// TIA Portal project "SSA-3GHz_V18" (V18)

(* hardware
DEVICE "S7-1200"  S7-1200 Station
   slot 0: "Stand.sectionalRail35mmLength483mm_0"  S7-1200 Rack  Rack  V1.0
   slot 1: "S7-1200"  CPU 1215C DC/DC/DC  6ES7 215-1AG40-0XB0  V4.5
   slot 2: "AnalogInputSM12314AI_2"  6ES7 231-4HD32-0XB0  V2.0
   slot 3: "S7-1200analogInputSM1231RTD4AI_3"  SM 1231 AI4 x RTD  6ES7 231-5PD32-0XB0  V2.0
DEVICE "HMI_1"  KTP400 Basic PN
   slot 0: "HMI_1"  KTP400 Basic PN  6AV2 123-2DB03-0AX0  15.1.0.0
   slot 1: "HMI_RT_1"  KTP400 Basic PN  6AV2 123-2DB03-0AX0  15.1.0.0
   slot 5: "HMI_1.IE_CP_1"  PROFINET Interface  15.0.1.0
      slot 1: "PROFINET Interface_1"  PROFINET Interface
         slot 1: "Port_1"  Port
*)

// ===== PLC "S7-1200"  CPU 1215C DC/DC/DC =====

VAR_GLOBAL   // PLC tag table "Default tag table"
   "System_Byte" AT %MB1 : Byte;
   "FirstScan" AT %M1.0 : Bool;
   "DiagStatusUpdate" AT %M1.1 : Bool;
   "AlwaysTRUE" AT %M1.2 : Bool;
   "AlwaysFALSE" AT %M1.3 : Bool;
   "Clock_Byte" AT %MB0 : Byte;
   "Clock_10Hz" AT %M0.0 : Bool;
   "Clock_5Hz" AT %M0.1 : Bool;
   "Clock_2.5Hz" AT %M0.2 : Bool;
   "Clock_2Hz" AT %M0.3 : Bool;
   "Clock_1.25Hz" AT %M0.4 : Bool;
   "Clock_1Hz" AT %M0.5 : Bool;
   "Clock_0.625Hz" AT %M0.6 : Bool;
   "Clock_0.5Hz" AT %M0.7 : Bool;
   "MoveBlkStat" AT %MW100 : Int;
   "tmp_setIP" AT %I1.1 : Bool;
   "Tag_2" AT %I1.2 : Bool;
   "Pulse_mem" AT %M10.1 : Bool;
   "Tag_3" AT %Q1.1 : Bool;
   "Modbus_srv_enable" AT %M2.3 : Bool;   // ModBus Server Enable bit
END_VAR

VAR_GLOBAL   // PLC tag table "Test tags"
   "Counter" AT %MD100 : UDInt;
   "TestBlink" AT %Q1.0 : Bool;
   "VisuTest" AT %MB104 : Byte;
   "Set_IP_PArameters" AT %M10.2 : Bool;
END_VAR

VAR_GLOBAL   // PLC tag table "Analog I/O"
   "U_drain_RBK" AT %IW64 : Int;   // Drain voltage read-back
   "U_drain" AT %QW64 : Int;   // Drain voltage set-point
   "ADC0ch1" AT %IW66 : Int;   // Spare
   "U_gate" AT %QW66 : Int;   // Gate voltage set-point
   "Pfwd" AT %IW96 : Int;   // Forward power
   "Prev" AT %IW98 : Int;   // Reverse power
   "I_drain" AT %IW100 : Int;   // Drain current
   "Pin" AT %IW102 : Int;   // Gate voltage read-back
   "TT01" AT %IW112 : Int;
   "TT02" AT %IW114 : Int;
   "TT03" AT %IW116 : Int;
   "TT04" AT %IW118 : Int;
END_VAR

VAR_GLOBAL   // PLC tag table "Digital I/O"
   "DutyCycOK" AT %I0.0 : Bool;   // Duty cycle OK
   "KeyIntlkOK" AT %I0.1 : Bool;   // Key interlock OK
   "ExtIntlk1" AT %I0.2 : Bool;   // DC PS enable
   "ExtIntlk2" AT %I0.3 : Bool;
   "T1_OK" AT %I0.4 : Bool;   // T1 trigger present
   "CoolingOK" AT %I0.5 : Bool;
   "Spare1" AT %I0.6 : Bool;   // Spare
   "FanOK" AT %I0.7 : Bool;   // Spare
   "ExtIntlkOK" AT %I1.0 : Bool;   // Spare
   "RFSwitchOn" AT %Q0.0 : Bool;   // Close RF switch
   "PSOutputOff" AT %Q0.1 : Bool;   // Set PS output off
   "SSA_OK" AT %Q0.2 : Bool;   // Solid State Amplifier OK - output interlock
   "ResetOut" AT %Q0.3 : Bool;   // Reset the errors signal out
   "cPSOn" AT %Q0.4 : Bool;   // When active 230 V AC is connected to the drain PS
END_VAR

VAR_GLOBAL   // PLC tag table "Memory tags"
   "RestoreFactorySettings" AT %M10.7 : Bool;   // Restore factory Settings (Ud look-up table and network settings)
END_VAR

TYPE "DigitalIN"
   STRUCT
      DigitalIN : Struct
         PhysIn : Bool;   // Physical input
         NegLogic : Bool;   // 0 - positive lgic, 1 - negative logic
         Disabled : Bool;   // 0 - signal enabled, 1 - signal disabled (not used in process controll)
         Out : Bool;   // Logical value after taking into accout NegLogic setting
      END_STRUCT;
   END_STRUCT;
END_TYPE

TYPE "AnalogOUT"
   STRUCT
      AnalogOUT : Struct
         In : Real;
         Out : Int;
         VisuState : Byte;
         MINDAC : Int;
         MAXDAC : Int;
         MINEGU : Real;
         MAXEGU : Real;
      END_STRUCT;
   END_STRUCT;
END_TYPE

TYPE "AnalogIN"
   STRUCT
      AnalogIN : Struct
         In : Word;
         Out : Real;
         Low : Real;
         LoLo : Real;
         High : Real;
         HIHi : Real;
         VisuState : Byte;
         MINADC : Int;
         MAXADC : Int;
         MINEGU : Real;
         MAXEGU : Real;
      END_STRUCT;
   END_STRUCT;
END_TYPE

TYPE "RTD_IN"
   STRUCT
      RTD_IN : Struct
         In : Word;
         Out : Real;
         Low : Real;
         LoLo : Real;
         High : Real;
         HIHi : Real;
         VisuState : Byte;
      END_STRUCT;
   END_STRUCT;
END_TYPE

DATA_BLOCK "IEC_Counter_0_DB"   // DB5
{ S7_Optimized_Access := 'TRUE' }
AUTHOR : Simatic
FAMILY : IEC
NAME : UDCNTR
VERSION : 1.2
// stored: InstanceOfName IEC_UDCOUNTER
"IEC_UDCOUNTER"
BEGIN
END_DATA_BLOCK

DATA_BLOCK "ModbusData"   // DB100
{ S7_Optimized_Access := 'TRUE' }
VERSION : 0.1
   VAR
      serverData : Struct
         disconnect : Bool;
         ndr : Bool;
         dataRead : Bool;
         error : Bool;
         status : Word;
         statusSave : Word;
      END_STRUCT;
   END_VAR
   VAR RETAIN
      connectParamServer : TCON_IP_v4;
   END_VAR
BEGIN
   connectParamServer.InterfaceId := 64;
   connectParamServer.ID := 16#1;
   connectParamServer.RemoteAddress.ADDR[1] := 0;
   connectParamServer.RemoteAddress.ADDR[2] := 0;
   connectParamServer.RemoteAddress.ADDR[3] := 0;
   connectParamServer.RemoteAddress.ADDR[4] := 0;
   connectParamServer.RemotePort := 0;
   connectParamServer.LocalPort := 502;
END_DATA_BLOCK

DATA_BLOCK "ModbusBuffer"   // DB101
{ S7_Optimized_Access := 'FALSE' }
VERSION : 0.1
   VAR
      BufferINOut : Struct
         LookupTable : Struct
            Pwr : Array[0..9] of Real;
            Ud : Array[0..9] of Real;
            Ug : Array[0..9] of Real;
         END_STRUCT;
         SetupData : Struct
            RemoteMode : Bool := FALSE;   // When true- remote control only
            dBm_unit : Bool := FALSE;   // When true - show power in dBm units
            NominalPower : Real := 100.0;   // Nominal Power
            NominalPower_dBm : Real := 50.0;   // Nominal Pwr [dBm]
            UdSP : Real := 17.91314;   // Udrain set-point
            UgSP : Real := 1.82;   // Ugate set-point
         END_STRUCT;
         Commands : Struct
            PSOutputOn : Bool := FALSE;
            PSOutputOff : Bool := FALSE;
            Stdby : Bool := FALSE;
            Reset : Bool := FALSE;
         END_STRUCT;
         ADCdata : Struct
            Udrain : Real := 0.0;
            Pin : Real := 0.0;
            Pfwd : Real := 0.0;
            Prev : Real := 0.0;
            Idrain : Real := 0.0;
            spare : Real := 0.0;
            TT01 : Real := 0.0;
            TT02 : Real := 0.0;
            TT03 : Real := 0.0;
            TT04 : Real := 0.0;
         END_STRUCT;
         CalculatedData : Struct
            Pfwd_dBm : Real := 0.0;
            Prev_dBm : Real := 0.0;
            Effic : Real;
            Pin_dBm : Real;
            AmplVisuState : Byte;
            spareByte : Byte;
            spare : Array[0..4] of Int;
         END_STRUCT;
         StatusBits : Struct
            DutyCycOK : Bool := FALSE;
            KeyIntlkOK : Bool := FALSE;
            ExtIntlk1 : Bool := FALSE;
            ExtIntlk2 : Bool := FALSE;
            T1_OK : Bool := FALSE;
            CoolingOK : Bool := FALSE;
            FanOK : Bool := FALSE;
            ExtIntlkOK : Bool := FALSE;
            DutyCycOK_Ign : Bool := FALSE;
            KeyIntlkOK_Ign : Bool := FALSE;
            ExtIntlk1_Ign : Bool := FALSE;
            ExtIntlk2_Ign : Bool := FALSE;
            T1_OK_Ign : Bool := FALSE;
            CoolingOK_Ign : Bool := TRUE;
            FanOK_Ign : Bool := FALSE;
            ExtIntlkOK_Ign : Bool := FALSE;
            RFSwitchON : Bool := FALSE;
            PSOutputOff : Bool;
            SSA_OK : Bool;
         END_STRUCT;
         Spare : Array[0..9] of Word;
         end : Word;
      END_STRUCT;
   END_VAR
BEGIN
   BufferINOut.LookupTable.Pwr[0] := 1.0;
   BufferINOut.LookupTable.Pwr[1] := 2.0;
   BufferINOut.LookupTable.Pwr[2] := 4.0;
   BufferINOut.LookupTable.Pwr[3] := 11.5;
   BufferINOut.LookupTable.Pwr[4] := 34.6;
   BufferINOut.LookupTable.Pwr[5] := 150.3;
   BufferINOut.LookupTable.Pwr[6] := 300.0;
   BufferINOut.LookupTable.Ud[0] := 13.5;
   BufferINOut.LookupTable.Ud[1] := 14.0;
   BufferINOut.LookupTable.Ud[2] := 14.5;
   BufferINOut.LookupTable.Ud[3] := 15.5;
   BufferINOut.LookupTable.Ud[4] := 16.5;
   BufferINOut.LookupTable.Ud[5] := 19.0;
   BufferINOut.LookupTable.Ud[6] := 23.5;
   BufferINOut.LookupTable.Ug[0] := 1.82;
   BufferINOut.LookupTable.Ug[1] := 1.82;
   BufferINOut.LookupTable.Ug[2] := 1.82;
   BufferINOut.LookupTable.Ug[3] := 1.82;
   BufferINOut.LookupTable.Ug[4] := 1.82;
   BufferINOut.LookupTable.Ug[5] := 1.82;
   BufferINOut.LookupTable.Ug[6] := 1.82;
   BufferINOut.LookupTable.Pwr[7] := 395.6;
   BufferINOut.LookupTable.Pwr[8] := 450.5;
   BufferINOut.LookupTable.Pwr[9] := 454.0;
   BufferINOut.LookupTable.Ud[7] := 27.5;
   BufferINOut.LookupTable.Ud[8] := 31.0;
   BufferINOut.LookupTable.Ud[9] := 32.0;
   BufferINOut.LookupTable.Ug[7] := 1.82;
   BufferINOut.LookupTable.Ug[8] := 1.82;
   BufferINOut.LookupTable.Ug[9] := 1.82;
   BufferINOut.CalculatedData.spare[0] := 0;
   BufferINOut.CalculatedData.spare[1] := 0;
   BufferINOut.CalculatedData.spare[2] := 0;
   BufferINOut.CalculatedData.spare[3] := 0;
END_DATA_BLOCK

DATA_BLOCK "HMIdata"   // DB103
{ S7_Optimized_Access := 'FALSE' }
VERSION : 0.1
   VAR
      Cordination : Word;
      getPlcMode : Int;
      plcTime : DTL;
      retValueTime : Word;
   END_VAR
BEGIN
END_DATA_BLOCK

DATA_BLOCK "DigitalInputs"   // DB400
{ S7_Optimized_Access := 'TRUE' }
VERSION : 0.1
   VAR
      DutyCycOK : "DigitalIN";
      KeyIntlkOK : "DigitalIN";
      ExtIntlk1 : "DigitalIN";
      ExtIntlk2 : "DigitalIN";
      T1_OK : "DigitalIN";
      CoolingOK : "DigitalIN";
      FanOK : "DigitalIN";   // Spare
      ExtIntlkOK : "DigitalIN";   // Spare
   END_VAR
BEGIN
   KeyIntlkOK.DigitalIN.Disabled := false;
   CoolingOK.DigitalIN.Disabled := false;
   FanOK.DigitalIN.Disabled := true;
   ExtIntlkOK.DigitalIN.Disabled := true;
   T1_OK.DigitalIN.Disabled := false;
END_DATA_BLOCK

DATA_BLOCK "AnalogInputs"   // DB401
{ S7_Optimized_Access := 'TRUE' }
VERSION : 0.1
   VAR
      U_drain_RBK : "AnalogIN";
      Pin : "AnalogIN";
      Pfwd : "AnalogIN";
      Prev : "AnalogIN";
      I_drain : "AnalogIN";
      ADC0ch1 : "AnalogIN";
      Pfwd_dBm : Real;
      Prev_dBm : Real;
      Pin_dBm : Real;
   END_VAR
   VAR RETAIN
      PinScale : Real := 3.0;
      PfwdScale : Real := 31.16;
      PrevScale : Real := 31.16;
   END_VAR
BEGIN
   U_drain_RBK.AnalogIN.MAXADC := 27648;
   Pin.AnalogIN.MINADC := 0;
   Pin.AnalogIN.MAXADC := 27648;
   Pfwd.AnalogIN.MAXADC := 27648;
   Pfwd.AnalogIN.MAXEGU := 67.6;
   Prev.AnalogIN.MAXADC := 27648;
   Prev.AnalogIN.MAXEGU := 62.1;
   I_drain.AnalogIN.MAXADC := 27648;
   I_drain.AnalogIN.MAXEGU := 15.0;
   ADC0ch1.AnalogIN.MAXADC := 27648;
   ADC0ch1.AnalogIN.MAXEGU := 10.0;
   U_drain_RBK.AnalogIN.MAXEGU := 48.0;
   Pin.AnalogIN.MAXEGU := 21.3;
   Pin.AnalogIN.MINEGU := -13.7;
   Pfwd.AnalogIN.MINEGU := 34.6;
   Prev.AnalogIN.MINEGU := 26.1;
END_DATA_BLOCK

DATA_BLOCK "AnalogOutputs"   // DB402
{ S7_Optimized_Access := 'TRUE' }
VERSION : 0.1
   VAR
      U_drain : "AnalogOUT";
      U_gate : "AnalogOUT";
   END_VAR
BEGIN
   U_drain.AnalogOUT.MAXDAC := 27648;
   U_drain.AnalogOUT.MAXEGU := 48.0;
   U_gate.AnalogOUT.MAXDAC := 27648;
   U_gate.AnalogOUT.MAXEGU := 5.0;
   U_gate.AnalogOUT.MINEGU := 0.0;
END_DATA_BLOCK

DATA_BLOCK "DigitalOutputs"   // DB450
{ S7_Optimized_Access := 'TRUE' }
VERSION : 0.1
   VAR
      RF_Switch_ON : Bool;
      ResetCmd : Bool;
      PSOutputOffCmd : Bool;
      PSOutputOnCmd : Bool;
      cPSOn : Bool;
   END_VAR
BEGIN
END_DATA_BLOCK

DATA_BLOCK "LookupTable"   // DB500
{ S7_Optimized_Access := 'FALSE' }
VERSION : 0.1
   VAR
      Pwr : Array[0..9] of Real;
      Ud : Array[0..9] of Real;
      Ug : Array[0..9] of Real;
   END_VAR
BEGIN
   Pwr[0] := 1.0;
   Pwr[1] := 2.0;
   Pwr[2] := 4.0;
   Pwr[3] := 11.5;
   Pwr[4] := 34.6;
   Pwr[5] := 150.3;
   Pwr[6] := 300.0;
   Ud[0] := 13.5;
   Ud[1] := 14.0;
   Ud[2] := 14.5;
   Ud[3] := 15.5;
   Ud[4] := 16.5;
   Ud[5] := 19.0;
   Ud[6] := 23.5;
   Ug[0] := 1.82;
   Ug[1] := 1.82;
   Ug[2] := 1.82;
   Ug[3] := 1.82;
   Ug[4] := 1.82;
   Ug[5] := 1.82;
   Ug[6] := 1.82;
   Pwr[7] := 395.6;
   Pwr[8] := 450.5;
   Pwr[9] := 454.0;
   Ud[7] := 27.5;
   Ud[8] := 31.0;
   Ud[9] := 32.0;
   Ug[7] := 1.82;
   Ug[8] := 1.82;
   Ug[9] := 1.82;
END_DATA_BLOCK

// folder: 5_T_CONFIG (S7-1200, S7-1500)

DATA_BLOCK "SLI_gDB_T_CONFIG_PLC"   // DB1
{ S7_Optimized_Access := 'TRUE' }
VERSION : 0.1
   VAR
      T_CONFIG : Struct   // Variables of T_CONFIG
         start : Bool;   // Set "start" to TRUE to configure the PROFINET interface.
         hwid : Hw_Interface := 64;   // Identification number of the PROFINET interface of the device (e. g. PROFINET interface of the CPU).
         busy : Bool;
         done : Bool;
         error : Bool;
         errorLocation : DWord;
         status : DWord;
         memErrStat : DWord;   // Saves the error status.
      END_STRUCT;
   END_VAR
   VAR RETAIN
      configData : Struct   // Data to configure the PROFINET device.
         header : IF_CONF_Header;   // The header is used to define the number of system data types.
         deviceIP : IF_CONF_v4;   // Specifies the IP of the PROFINET device.
         deviceName : IF_CONF_NOS;   // Specifies the name of the PROFINET interface ("PROFINET device name").
      END_STRUCT;
   END_VAR
BEGIN
   configData.header.SubfieldCount := 2;   // 2: Indicates that two additional structures ("deviceIP" and "deviceName") are used below.
   configData.deviceName.Length := 11;   // Information on overall length of the structure (5 bytes for the device name "myplc" + 6 bytes for the parameters Id, Length and Mode)
   configData.deviceName.Mode := 1;   // 1: Permanent change of the device name in "myplc".
   configData.deviceName.NOS[1] := 'm';
   configData.deviceName.NOS[2] := 'y';
   configData.deviceName.NOS[3] := 'p';
   configData.deviceName.NOS[4] := 'l';
   configData.deviceName.NOS[5] := 'c';
   configData.deviceIP.Length := 18;   // Information on overall length of the structure (12 bytes for the device IP + 6 bytes for the parameters Id, Length and Mode)
   configData.deviceIP.Mode := 1;   // 1: Permanent change of the device IP.
   configData.deviceIP.InterfaceAddress.ADDR[1] := 192;
   configData.deviceIP.InterfaceAddress.ADDR[2] := 168;
   configData.deviceIP.InterfaceAddress.ADDR[3] := 1;
   configData.deviceIP.InterfaceAddress.ADDR[4] := 234;
   configData.deviceIP.SubnetMask.ADDR[1] := 255;
   configData.deviceIP.SubnetMask.ADDR[2] := 255;
   configData.deviceIP.SubnetMask.ADDR[3] := 255;
   configData.deviceIP.SubnetMask.ADDR[4] := 0;
   configData.deviceIP.DefaultRouter.ADDR[1] := 192;
   configData.deviceIP.DefaultRouter.ADDR[2] := 168;
   configData.deviceIP.DefaultRouter.ADDR[3] := 1;
   configData.deviceIP.DefaultRouter.ADDR[4] := 1;
   // configData.header.FieldType : Field type: Must always have the value "0".
   // configData.header.FieldId : Error ID: Must always have the value "0".
   // configData.deviceIP.Id : System data type ID. The start value of this parameter must not be changed.
   // configData.deviceIP.InterfaceAddress : IP connection data. IP address
   // configData.deviceIP.SubnetMask : IP connection data. Subnet mask
   // configData.deviceIP.DefaultRouter : IP connection data. Router address (optional)
   // configData.deviceName.Id : System data type ID. The start value of this parameter must not be changed.
   // configData.deviceName.NOS : Device name (1 character per byte)
END_DATA_BLOCK

// folder: System blocks/Program resources

DATA_BLOCK "IEC_Timer_0_DB"   // DB6
{ S7_Optimized_Access := 'TRUE' }
AUTHOR : Simatic
FAMILY : IEC
NAME : IEC_TMR
VERSION : 1.0
// stored: InstanceOfName IEC_TIMER
"IEC_TIMER"
BEGIN
END_DATA_BLOCK

DATA_BLOCK "ResetCmdTimer"   // DB7
{ S7_Optimized_Access := 'TRUE' }
AUTHOR : Simatic
FAMILY : IEC
NAME : IEC_TMR
VERSION : 1.0
// stored: InstanceOfName IEC_TIMER
"IEC_TIMER"
BEGIN
END_DATA_BLOCK

// folder: (top level)

FUNCTION "Tests" : Void   // FC1, LAD
{ S7_Optimized_Access := 'TRUE' }
VERSION : 0.1
BEGIN

REGION Network 1
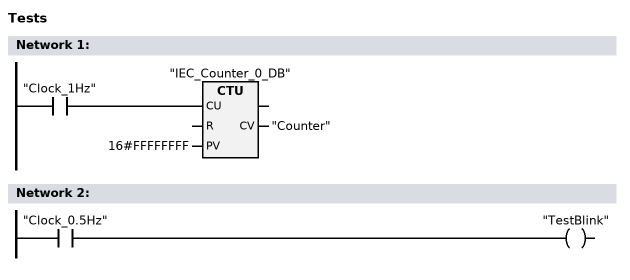
   "IEC_Counter_0_DB".CTU(CU := "Clock_1Hz", PV := 16#FFFFFFFF, CV => "Counter");
END_REGION

REGION Network 2
   RUNG wire#powerrail
      Contact( "Clock_0.5Hz" )
      Coil( "TestBlink" )
   END_RUNG
   // the same network as SCL:
   "TestBlink" := "Clock_0.5Hz";
END_REGION
END_FUNCTION

FUNCTION "ScalePowerADC" : Void   // FC2, SCL
{ S7_Optimized_Access := 'TRUE' }
VERSION : 0.1
   VAR_INPUT
      InData : Word;
   END_VAR
   VAR_OUTPUT
      Pwr_dBm : Real;
   END_VAR
   VAR_IN_OUT
      AInp : "AnalogIN";   // Analog Input structure
   END_VAR
   VAR_TEMP
      tmpR : Real;
   END_VAR
   VAR CONSTANT
      LN_10 : Real := 2.302585;   // ln(10)
   END_VAR
BEGIN
   REGION LinearScaling
       // Statement section REGION
       #AInp.AnalogIN.In := #InData;
       #tmpR := NORM_X(MIN := #AInp.AnalogIN.MINADC, VALUE := #AInp.AnalogIN.In, MAX := #AInp.AnalogIN.MAXADC);
       #Pwr_dBm := SCALE_X(MIN := #AInp.AnalogIN.MINEGU, VALUE := #tmpR, MAX := #AInp.AnalogIN.MAXEGU);
   END_REGION
   REGION Convertion_to_W
       // Statement section REGION
       #tmpR := #LN_10 * #Pwr_dBm / 10;
       #AInp.AnalogIN.Out := EXP(#tmpR) / 1000;
   END_REGION
END_FUNCTION

FUNCTION "Modbus2PLC" : Void   // FC10, LAD
{ S7_Optimized_Access := 'TRUE' }
VERSION : 0.1
   VAR_TEMP   // added for the SCL form of the ladder/FBD networks
      _w1 : Bool;
   END_VAR
BEGIN

REGION Network 1: Save the current look-up table to the factory settings table
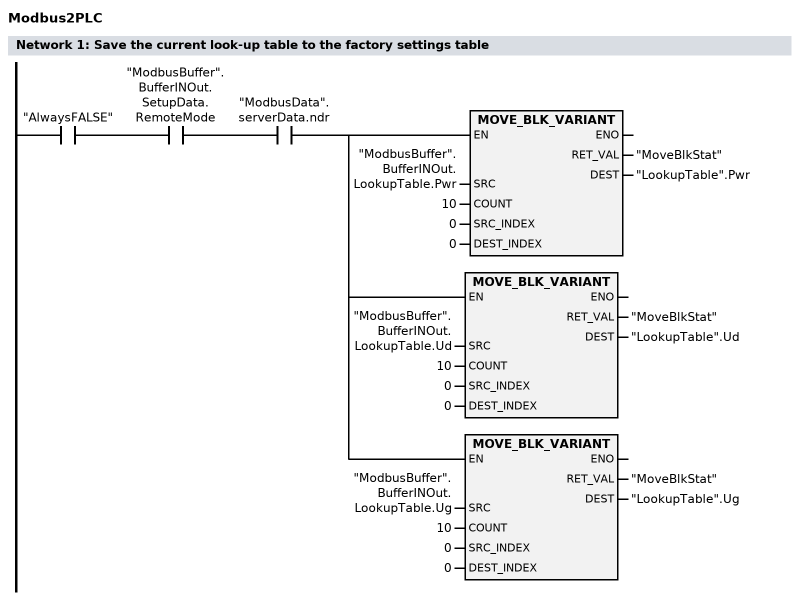
   #_w1 := "AlwaysFALSE" AND "ModbusBuffer".BufferINOut.SetupData.RemoteMode AND "ModbusData".serverData.ndr;
   IF #_w1 THEN
       "MoveBlkStat" := MOVE_BLK_VARIANT(SRC := "ModbusBuffer".BufferINOut.LookupTable.Pwr,
                               COUNT := 10,
                               SRC_INDEX := 0,
                               DEST_INDEX := 0,
                               DEST => "LookupTable".Pwr);
       "MoveBlkStat" := MOVE_BLK_VARIANT(SRC := "ModbusBuffer".BufferINOut.LookupTable.Ud,
                               COUNT := 10,
                               SRC_INDEX := 0,
                               DEST_INDEX := 0,
                               DEST => "LookupTable".Ud);
       "MoveBlkStat" := MOVE_BLK_VARIANT(SRC := "ModbusBuffer".BufferINOut.LookupTable.Ug,
                               COUNT := 10,
                               SRC_INDEX := 0,
                               DEST_INDEX := 0,
                               DEST => "LookupTable".Ug);
   END_IF;
END_REGION
END_FUNCTION

FUNCTION "PLC2Modbus" : Void   // FC11, LAD
{ S7_Optimized_Access := 'TRUE' }
VERSION : 0.1
   VAR_TEMP   // added for the SCL form of the ladder/FBD networks
      _w1 : Bool;
   END_VAR
BEGIN

REGION Network 1: Restore the factory settings
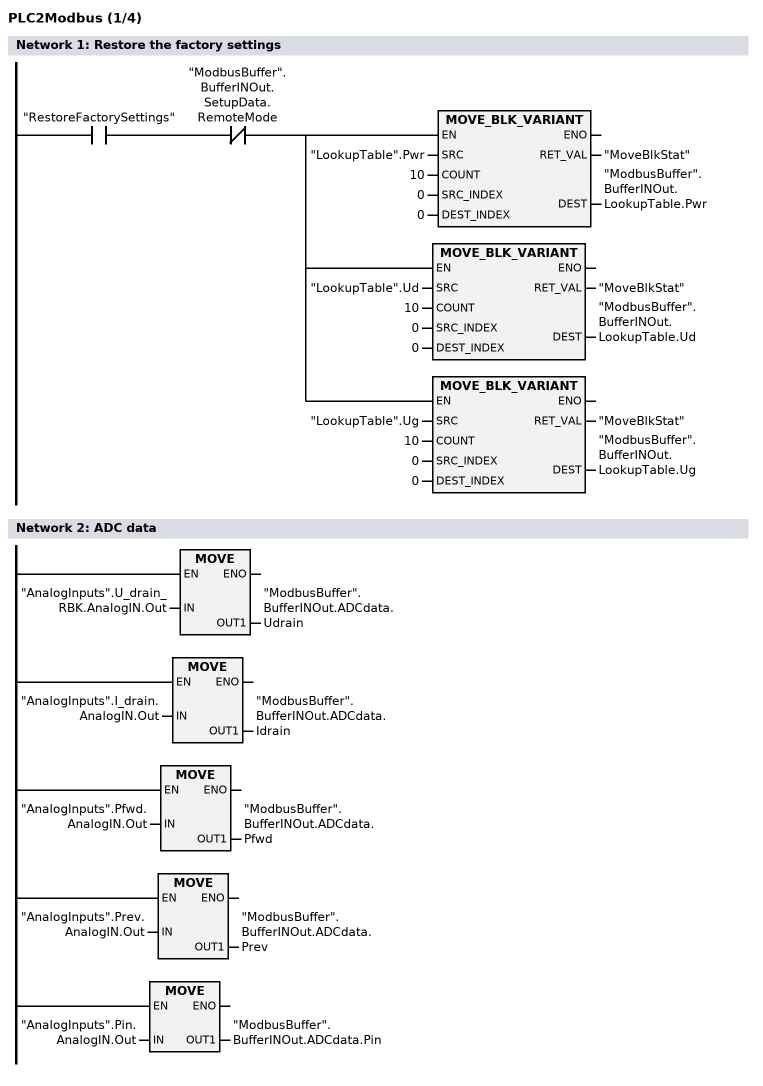
   #_w1 := "RestoreFactorySettings" AND NOT "ModbusBuffer".BufferINOut.SetupData.RemoteMode;
   IF #_w1 THEN
       "MoveBlkStat" := MOVE_BLK_VARIANT(SRC := "LookupTable".Pwr,
                               COUNT := 10,
                               SRC_INDEX := 0,
                               DEST_INDEX := 0,
                               DEST => "ModbusBuffer".BufferINOut.LookupTable.Pwr);
       "MoveBlkStat" := MOVE_BLK_VARIANT(SRC := "LookupTable".Ud,
                               COUNT := 10,
                               SRC_INDEX := 0,
                               DEST_INDEX := 0,
                               DEST => "ModbusBuffer".BufferINOut.LookupTable.Ud);
       "MoveBlkStat" := MOVE_BLK_VARIANT(SRC := "LookupTable".Ug,
                               COUNT := 10,
                               SRC_INDEX := 0,
                               DEST_INDEX := 0,
                               DEST => "ModbusBuffer".BufferINOut.LookupTable.Ug);
   END_IF;
END_REGION

REGION Network 2: ADC data
   RUNG wire#powerrail
      Move(in := "AnalogInputs".U_drain_RBK.AnalogIN.Out, out1 => "ModbusBuffer".BufferINOut.ADCdata.Udrain)
   END_RUNG
   RUNG wire#powerrail
      Move(in := "AnalogInputs".I_drain.AnalogIN.Out, out1 => "ModbusBuffer".BufferINOut.ADCdata.Idrain)
   END_RUNG
   RUNG wire#powerrail
      Move(in := "AnalogInputs".Pfwd.AnalogIN.Out, out1 => "ModbusBuffer".BufferINOut.ADCdata.Pfwd)
   END_RUNG
   RUNG wire#powerrail
      Move(in := "AnalogInputs".Prev.AnalogIN.Out, out1 => "ModbusBuffer".BufferINOut.ADCdata.Prev)
   END_RUNG
   RUNG wire#powerrail
      Move(in := "AnalogInputs".Pin.AnalogIN.Out, out1 => "ModbusBuffer".BufferINOut.ADCdata.Pin)
   END_RUNG
   // the same network as SCL:
   "ModbusBuffer".BufferINOut.ADCdata.Udrain := "AnalogInputs".U_drain_RBK.AnalogIN.Out;
   "ModbusBuffer".BufferINOut.ADCdata.Idrain := "AnalogInputs".I_drain.AnalogIN.Out;
   "ModbusBuffer".BufferINOut.ADCdata.Pfwd := "AnalogInputs".Pfwd.AnalogIN.Out;
   "ModbusBuffer".BufferINOut.ADCdata.Prev := "AnalogInputs".Prev.AnalogIN.Out;
   "ModbusBuffer".BufferINOut.ADCdata.Pin := "AnalogInputs".Pin.AnalogIN.Out;
END_REGION

REGION Network 3: Calculated data
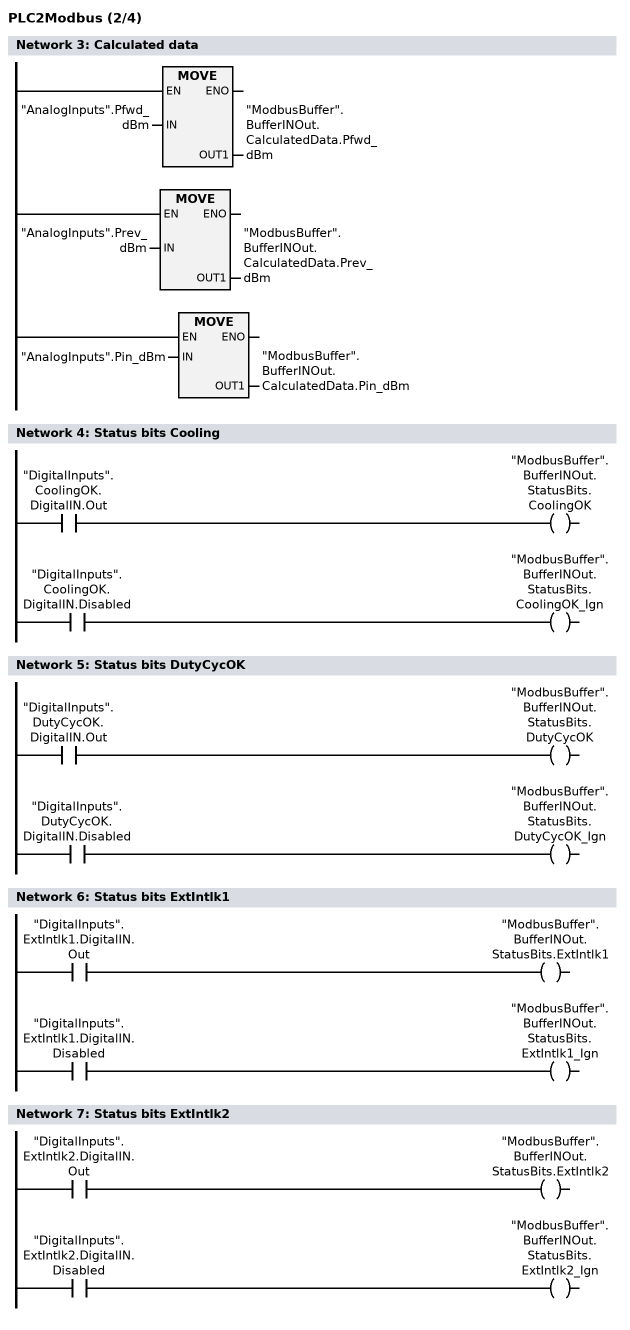
   RUNG wire#powerrail
      Move(in := "AnalogInputs".Pfwd_dBm, out1 => "ModbusBuffer".BufferINOut.CalculatedData.Pfwd_dBm)
   END_RUNG
   RUNG wire#powerrail
      Move(in := "AnalogInputs".Prev_dBm, out1 => "ModbusBuffer".BufferINOut.CalculatedData.Prev_dBm)
   END_RUNG
   RUNG wire#powerrail
      Move(in := "AnalogInputs".Pin_dBm, out1 => "ModbusBuffer".BufferINOut.CalculatedData.Pin_dBm)
   END_RUNG
   // the same network as SCL:
   "ModbusBuffer".BufferINOut.CalculatedData.Pfwd_dBm := "AnalogInputs".Pfwd_dBm;
   "ModbusBuffer".BufferINOut.CalculatedData.Prev_dBm := "AnalogInputs".Prev_dBm;
   "ModbusBuffer".BufferINOut.CalculatedData.Pin_dBm := "AnalogInputs".Pin_dBm;
END_REGION

REGION Network 4: Status bits Cooling
   RUNG wire#powerrail
      Contact( "DigitalInputs".CoolingOK.DigitalIN.Out )
      Coil( "ModbusBuffer".BufferINOut.StatusBits.CoolingOK )
   END_RUNG
   RUNG wire#powerrail
      Contact( "DigitalInputs".CoolingOK.DigitalIN.Disabled )
      Coil( "ModbusBuffer".BufferINOut.StatusBits.CoolingOK_Ign )
   END_RUNG
   // the same network as SCL:
   "ModbusBuffer".BufferINOut.StatusBits.CoolingOK := "DigitalInputs".CoolingOK.DigitalIN.Out;
   "ModbusBuffer".BufferINOut.StatusBits.CoolingOK_Ign := "DigitalInputs".CoolingOK.DigitalIN.Disabled;
END_REGION

REGION Network 5: Status bits DutyCycOK
   RUNG wire#powerrail
      Contact( "DigitalInputs".DutyCycOK.DigitalIN.Out )
      Coil( "ModbusBuffer".BufferINOut.StatusBits.DutyCycOK )
   END_RUNG
   RUNG wire#powerrail
      Contact( "DigitalInputs".DutyCycOK.DigitalIN.Disabled )
      Coil( "ModbusBuffer".BufferINOut.StatusBits.DutyCycOK_Ign )
   END_RUNG
   // the same network as SCL:
   "ModbusBuffer".BufferINOut.StatusBits.DutyCycOK := "DigitalInputs".DutyCycOK.DigitalIN.Out;
   "ModbusBuffer".BufferINOut.StatusBits.DutyCycOK_Ign := "DigitalInputs".DutyCycOK.DigitalIN.Disabled;
END_REGION

REGION Network 6: Status bits ExtIntlk1
   RUNG wire#powerrail
      Contact( "DigitalInputs".ExtIntlk1.DigitalIN.Out )
      Coil( "ModbusBuffer".BufferINOut.StatusBits.ExtIntlk1 )
   END_RUNG
   RUNG wire#powerrail
      Contact( "DigitalInputs".ExtIntlk1.DigitalIN.Disabled )
      Coil( "ModbusBuffer".BufferINOut.StatusBits.ExtIntlk1_Ign )
   END_RUNG
   // the same network as SCL:
   "ModbusBuffer".BufferINOut.StatusBits.ExtIntlk1 := "DigitalInputs".ExtIntlk1.DigitalIN.Out;
   "ModbusBuffer".BufferINOut.StatusBits.ExtIntlk1_Ign := "DigitalInputs".ExtIntlk1.DigitalIN.Disabled;
END_REGION

REGION Network 7: Status bits ExtIntlk2
   RUNG wire#powerrail
      Contact( "DigitalInputs".ExtIntlk2.DigitalIN.Out )
      Coil( "ModbusBuffer".BufferINOut.StatusBits.ExtIntlk2 )
   END_RUNG
   RUNG wire#powerrail
      Contact( "DigitalInputs".ExtIntlk2.DigitalIN.Disabled )
      Coil( "ModbusBuffer".BufferINOut.StatusBits.ExtIntlk2_Ign )
   END_RUNG
   // the same network as SCL:
   "ModbusBuffer".BufferINOut.StatusBits.ExtIntlk2 := "DigitalInputs".ExtIntlk2.DigitalIN.Out;
   "ModbusBuffer".BufferINOut.StatusBits.ExtIntlk2_Ign := "DigitalInputs".ExtIntlk2.DigitalIN.Disabled;
END_REGION

REGION Network 8: Status bits KeyIntlkOK
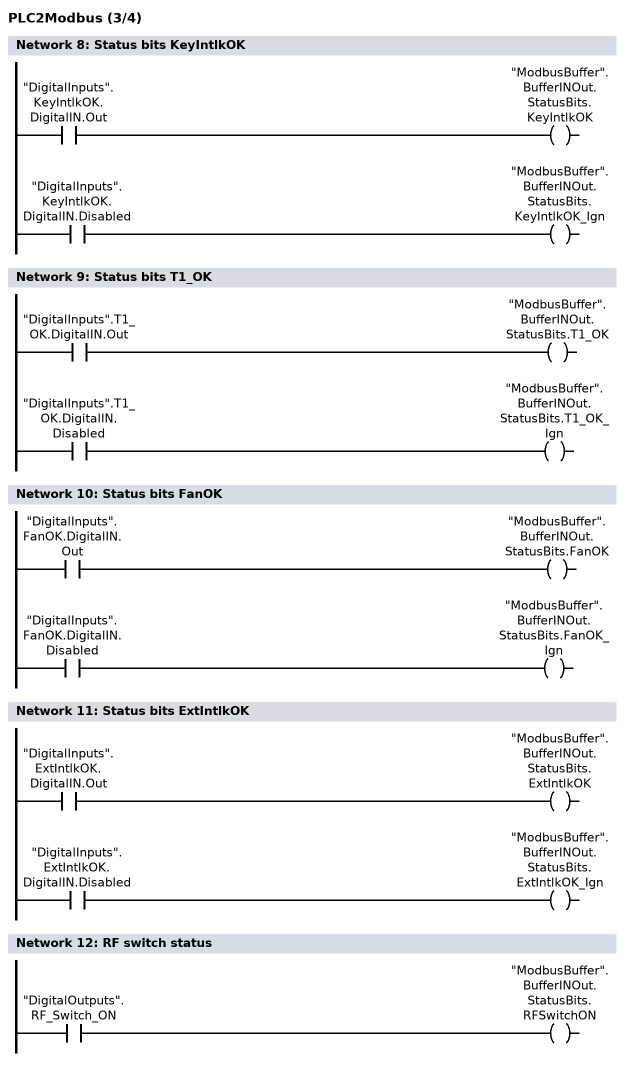
   RUNG wire#powerrail
      Contact( "DigitalInputs".KeyIntlkOK.DigitalIN.Out )
      Coil( "ModbusBuffer".BufferINOut.StatusBits.KeyIntlkOK )
   END_RUNG
   RUNG wire#powerrail
      Contact( "DigitalInputs".KeyIntlkOK.DigitalIN.Disabled )
      Coil( "ModbusBuffer".BufferINOut.StatusBits.KeyIntlkOK_Ign )
   END_RUNG
   // the same network as SCL:
   "ModbusBuffer".BufferINOut.StatusBits.KeyIntlkOK := "DigitalInputs".KeyIntlkOK.DigitalIN.Out;
   "ModbusBuffer".BufferINOut.StatusBits.KeyIntlkOK_Ign := "DigitalInputs".KeyIntlkOK.DigitalIN.Disabled;
END_REGION

REGION Network 9: Status bits T1_OK
   RUNG wire#powerrail
      Contact( "DigitalInputs".T1_OK.DigitalIN.Out )
      Coil( "ModbusBuffer".BufferINOut.StatusBits.T1_OK )
   END_RUNG
   RUNG wire#powerrail
      Contact( "DigitalInputs".T1_OK.DigitalIN.Disabled )
      Coil( "ModbusBuffer".BufferINOut.StatusBits.T1_OK_Ign )
   END_RUNG
   // the same network as SCL:
   "ModbusBuffer".BufferINOut.StatusBits.T1_OK := "DigitalInputs".T1_OK.DigitalIN.Out;
   "ModbusBuffer".BufferINOut.StatusBits.T1_OK_Ign := "DigitalInputs".T1_OK.DigitalIN.Disabled;
END_REGION

REGION Network 10: Status bits FanOK
   RUNG wire#powerrail
      Contact( "DigitalInputs".FanOK.DigitalIN.Out )
      Coil( "ModbusBuffer".BufferINOut.StatusBits.FanOK )
   END_RUNG
   RUNG wire#powerrail
      Contact( "DigitalInputs".FanOK.DigitalIN.Disabled )
      Coil( "ModbusBuffer".BufferINOut.StatusBits.FanOK_Ign )
   END_RUNG
   // the same network as SCL:
   "ModbusBuffer".BufferINOut.StatusBits.FanOK := "DigitalInputs".FanOK.DigitalIN.Out;
   "ModbusBuffer".BufferINOut.StatusBits.FanOK_Ign := "DigitalInputs".FanOK.DigitalIN.Disabled;
END_REGION

REGION Network 11: Status bits ExtIntlkOK
   RUNG wire#powerrail
      Contact( "DigitalInputs".ExtIntlkOK.DigitalIN.Out )
      Coil( "ModbusBuffer".BufferINOut.StatusBits.ExtIntlkOK )
   END_RUNG
   RUNG wire#powerrail
      Contact( "DigitalInputs".ExtIntlkOK.DigitalIN.Disabled )
      Coil( "ModbusBuffer".BufferINOut.StatusBits.ExtIntlkOK_Ign )
   END_RUNG
   // the same network as SCL:
   "ModbusBuffer".BufferINOut.StatusBits.ExtIntlkOK := "DigitalInputs".ExtIntlkOK.DigitalIN.Out;
   "ModbusBuffer".BufferINOut.StatusBits.ExtIntlkOK_Ign := "DigitalInputs".ExtIntlkOK.DigitalIN.Disabled;
END_REGION

REGION Network 12: RF switch status
   RUNG wire#powerrail
      Contact( "DigitalOutputs".RF_Switch_ON )
      Coil( "ModbusBuffer".BufferINOut.StatusBits.RFSwitchON )
   END_RUNG
   // the same network as SCL:
   "ModbusBuffer".BufferINOut.StatusBits.RFSwitchON := "DigitalOutputs".RF_Switch_ON;
END_REGION

REGION Network 13: Amplifier visual state
   // Calculates the enum vallue for the amplidier's visual state:
   // state 1 (blue): 230 V to drain PS connected, PS output off
   // state 2 (green): 230 V to drain PS connected, PS output on
   // state 4 (red): 230 V to drain PS disconnected
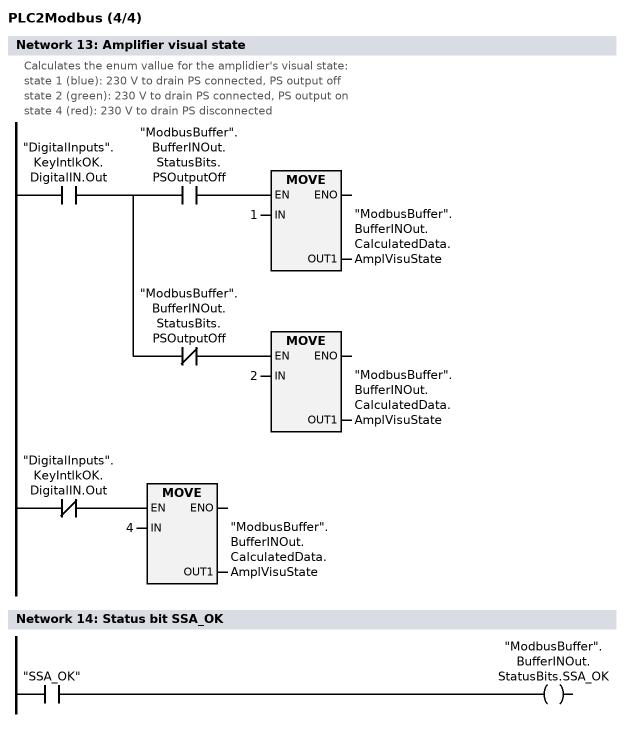
   RUNG wire#powerrail
      Contact( "DigitalInputs".KeyIntlkOK.DigitalIN.Out )
      wire#w1
      Contact( "ModbusBuffer".BufferINOut.StatusBits.PSOutputOff )
      Move(in := 1, out1 => "ModbusBuffer".BufferINOut.CalculatedData.AmplVisuState)
   END_RUNG
   RUNG wire#w1
      I_Contact( "ModbusBuffer".BufferINOut.StatusBits.PSOutputOff )
      Move(in := 2, out1 => "ModbusBuffer".BufferINOut.CalculatedData.AmplVisuState)
   END_RUNG
   RUNG wire#powerrail
      I_Contact( "DigitalInputs".KeyIntlkOK.DigitalIN.Out )
      Move(in := 4, out1 => "ModbusBuffer".BufferINOut.CalculatedData.AmplVisuState)
   END_RUNG
   // the same network as SCL:
   IF "DigitalInputs".KeyIntlkOK.DigitalIN.Out AND "ModbusBuffer".BufferINOut.StatusBits.PSOutputOff THEN
       "ModbusBuffer".BufferINOut.CalculatedData.AmplVisuState := 1;
   END_IF;
   IF "DigitalInputs".KeyIntlkOK.DigitalIN.Out AND NOT "ModbusBuffer".BufferINOut.StatusBits.PSOutputOff THEN
       "ModbusBuffer".BufferINOut.CalculatedData.AmplVisuState := 2;
   END_IF;
   IF NOT "DigitalInputs".KeyIntlkOK.DigitalIN.Out THEN
       "ModbusBuffer".BufferINOut.CalculatedData.AmplVisuState := 4;
   END_IF;
END_REGION

REGION Network 14: Status bit SSA_OK
   RUNG wire#powerrail
      Contact( "SSA_OK" )
      Coil( "ModbusBuffer".BufferINOut.StatusBits.SSA_OK )
   END_RUNG
   // the same network as SCL:
   "ModbusBuffer".BufferINOut.StatusBits.SSA_OK := "SSA_OK";
END_REGION
END_FUNCTION

FUNCTION "Setup" : Void   // FC90, LAD
{ S7_Optimized_Access := 'TRUE' }
VERSION : 0.1
// Set-up PROFINET interfaces.
   VAR_TEMP
      done_PLC : Bool;
      done_HMI : Bool;
      errorLocation_PLC : DWord;
      errorLocation_HMI : DWord;
   END_VAR
   VAR_TEMP   // added for the SCL form of the ladder/FBD networks
      _w1 : Bool;
      _w2 : Bool;
   END_VAR
BEGIN

REGION Network 1: Restore the factory setting for the network interface